// TIA Portal project "UploadAG314C_tia" (V15)

(* hardware
DEVICE "SIMATIC 300(1)"  S7-300 station
   slot 0: "Rack 0"  Rail  6ES7 390-1***0-0AA0
   slot 2: "CPU 314C-2 DP"  CPU 314C-2 DP  6ES7 314-6CG03-0AB0  V2.6
      slot 0: "MPI interface_1"  X1
      slot 1: "DP interface_1"  X2
      slot 2: "DI 24/DO 16_1"  DI24/DO16
      slot 3: "AI 5/AO 2_1"  AI5/AO2
      slot 4: "Count_1"  Counter
      slot 5: "Positioning_1"  Positioning
DEVICE "Test_Pump"  TP1200 Comfort
   slot 0: "Test_Pump"  TP1200 Comfort  6AV2 124-0MC01-0AX0  14.0.1.0
   slot 1: "HMI_RT_2"  TP1200 Comfort  6AV2 124-0MC01-0AX0  14.0.1.0
   slot 5: "Test_Pump._CP_1"  PROFINET Interface  14.0.1.0
      slot 1: "PROFINET Interface_1"  PROFINET Interface
         slot 1: "Port_1"  Port
         slot 2: "Port_2"  Port
   slot 7: "Test_Pump.I/DP_CP_1"  MPI/DP Interface  14.0.1.0
*)

// ===== PLC "CPU 314C-2 DP"  CPU 314C-2 DP =====
// protected blocks, not shown: "CONT_C_LF"

VAR_GLOBAL   // PLC tag table "Default tag table"
   "Tag_5" AT %M40.0 : Bool;
   "Tag_6" AT %M30.0 : Bool;
   "Tag_7" AT %M30.3 : Bool;
   "Tag_8" AT %M30.6 : Bool;
   "Tag_9" AT %M30.4 : Bool;
   "Tag_10" AT %M30.7 : Bool;
   "Tag_11" AT %M33.3 : Bool;
   "Tag_12" AT %M33.6 : Bool;
   "Tag_13" AT %M33.4 : Bool;
   "Tag_14" AT %M33.7 : Bool;
   "Tag_15" AT %I126.0 : Bool;
   "Tag_16" AT %M70.1 : Bool;
   "Tag_17" AT %I126.1 : Bool;
   "Tag_18" AT %M70.0 : Bool;
   "Tag_19" AT %I126.2 : Bool;
   "Tag_20" AT %I126.3 : Bool;
   "Tag_21" AT %I126.5 : Bool;
   "Tag_22" AT %I126.6 : Bool;
   "Tag_23" AT %Q124.1 : Bool;
   "Tag_24" AT %Q124.0 : Bool;
   "Tag_25" AT %M30.1 : Bool;
   "Tag_26" AT %M31.0 : Bool;
   "Tag_27" AT %T40 : Timer;
   "Tag_28" AT %Q124.2 : Bool;
   "Tag_29" AT %MD210 : DWord;
   "Tag_30" AT %MW212 : Word;
   "samplingTimer_1" AT %T190 : Timer;
   "samplingTimer_2" AT %T191 : Timer;
   "Tag_31" AT %M0.0 : Bool;
   "Tag_32" AT %T192 : Timer;
   "Speed" AT %MW4 : Int;
END_VAR

VAR_GLOBAL   // PLC tag table "STEP7 classic symbols"
   "Tag_1" AT %AW752 : Word;
   "Tag_2" AT %EW752 : Int;
   "Tag_3" AT %EW760 : Word;
   "Tag_4" AT %MD20 : DInt;
END_VAR

DATA_BLOCK "DB3"   // DB3
{ S7_Optimized_Access := 'FALSE' }
VERSION : 0.1
   VAR
      STAT0 : Word := WORD#16#0001;
      STAT1 : Word;
      STAT2 : Word := WORD#16#0009;
      STAT3 : Word := WORD#16#0003;
      STAT4 : Word := WORD#16#0027;
      STAT5 : Word := WORD#16#1456;
      STAT6 : Word;
      STAT7 : Word;
      STAT8 : Word;
      STAT9 : Word;
      STAT10 : Word;
      STAT11 : Word;
      STAT12 : Word;
      STAT13 : Word;
      STAT14 : Word;
      STAT15 : Word;
      STAT16 : Word;
      STAT17 : Word;
      STAT18 : Word;
      STAT19 : Word;
      STAT20 : Word;
   END_VAR
BEGIN
END_DATA_BLOCK

DATA_BLOCK "DB5"   // DB5
{ S7_Optimized_Access := 'FALSE' }
VERSION : 0.1
   VAR
      STAT0 : Word;
      STAT1 : Word := WORD#16#0400;
      STAT2 : Word;
      STAT3 : Word := WORD#16#0001;
      STAT4 : Word := WORD#16#0001;
      STAT5 : Word := WORD#16#0020;
      STAT6 : Word;
      STAT7 : Word;
      STAT8 : Word;
      STAT9 : Word;
      STAT10 : Word;
      STAT11 : Word;
      STAT12 : Word;
      STAT13 : Word;
      STAT14 : Word;
      STAT15 : Word;
      STAT16 : Word;
      STAT17 : Word;
      STAT18 : Word;
      STAT19 : Word;
      STAT20 : Word;
   END_VAR
BEGIN
END_DATA_BLOCK

DATA_BLOCK "DB12"   // DB12
{ S7_Optimized_Access := 'FALSE' }
VERSION : 0.1
   VAR
      STAT0 : Int;
      STAT1 : Int;
      STAT2 : Int := 250;
      STAT3 : Int := 336;
      STAT4 : DInt;
      STAT5 : DInt;
      STAT6 : DInt;
      STAT7 : DInt;
      STAT8 : DInt;
      STAT9 : DInt;
      STAT10 : DInt;
   END_VAR
BEGIN
END_DATA_BLOCK

DATA_BLOCK "DB13"   // DB13
{ S7_Optimized_Access := 'FALSE' }
VERSION : 0.1
   VAR
      STAT0 : Real;
      STAT1 : Real;
      STAT2 : Real;
      STAT3 : Real;
      STAT4 : Real;
      STAT5 : Real;
      STAT6 : Real;
      STAT7 : Real;
   END_VAR
BEGIN
END_DATA_BLOCK

DATA_BLOCK "DB14"   // DB14
{ S7_Optimized_Access := 'FALSE' }
VERSION : 0.1
   VAR
      STAT0 : Int;
      STAT1 : Int;
      STAT2 : DInt;
      STAT3 : DInt;
      STAT4 : DInt;
      STAT5 : Int;
      STAT6 : Int;
      STAT7 : Int := 410;
      STAT8 : Int;
      STAT9 : DInt;
      STAT10 : DInt;
      STAT11 : DInt;
      STAT12 : Int := 6800;
      STAT13 : Int;
      STAT14 : DInt;
      STAT15 : DInt;
      STAT16 : DInt;
      STAT17 : DInt;
      STAT18 : Real;
      STAT19 : Real;
      STAT20 : DInt;
      STAT21 : DInt := DINT#98300;
      STAT22 : Real;
      STAT23 : Real;
      STAT24 : Real;
   END_VAR
BEGIN
END_DATA_BLOCK

DATA_BLOCK "DB16"   // DB16
{ S7_Optimized_Access := 'FALSE' }
VERSION : 0.1
   VAR
      STAT0 : Int;
      STAT1 : String[10];
      STAT2 : DInt;
      STAT3 : DInt;
      STAT4 : DInt;
      STAT5 : DInt := DINT#750;
      STAT6 : DInt;
      STAT7 : DInt;
      STAT8 : DInt;
      STAT9 : DInt;
      STAT10 : DInt;
      STAT11 : DInt;
      STAT12 : DInt;
      STAT13 : Int;
      STAT14 : Int := 1;
      STAT15 : String[10];
      STAT16 : DInt;
      STAT17 : DInt;
      STAT18 : DInt;
      STAT19 : DInt;
      STAT20 : DInt;
      STAT21 : DInt;
      STAT22 : DInt;
      STAT23 : DInt;
      STAT24 : DInt;
      STAT25 : DInt;
      STAT26 : DInt;
      STAT27 : Int;
      STAT28 : Int := 2;
      STAT29 : String[10];
      STAT30 : DInt;
      STAT31 : DInt;
      STAT32 : DInt;
      STAT33 : DInt;
      STAT34 : DInt;
      STAT35 : DInt;
      STAT36 : DInt;
      STAT37 : DInt;
      STAT38 : DInt;
      STAT39 : DInt;
      STAT40 : DInt;
      STAT41 : Int;
      STAT42 : Int := 3;
      STAT43 : String[10];
      STAT44 : DInt;
      STAT45 : DInt;
      STAT46 : DInt;
      STAT47 : DInt;
      STAT48 : DInt;
      STAT49 : DInt;
      STAT50 : DInt;
      STAT51 : DInt;
      STAT52 : DInt;
      STAT53 : DInt;
      STAT54 : DInt;
      STAT55 : Int;
      STAT56 : Int := 4;
      STAT57 : String[10];
      STAT58 : DInt;
      STAT59 : DInt;
      STAT60 : DInt;
      STAT61 : DInt;
      STAT62 : DInt;
      STAT63 : DInt;
      STAT64 : DInt;
      STAT65 : DInt;
      STAT66 : DInt;
      STAT67 : DInt;
      STAT68 : DInt;
      STAT69 : Int;
      STAT70 : Int := 5;
      STAT71 : String[10];
      STAT72 : DInt;
      STAT73 : DInt;
      STAT74 : DInt;
      STAT75 : DInt;
      STAT76 : DInt;
      STAT77 : DInt;
      STAT78 : DInt;
      STAT79 : DInt;
      STAT80 : DInt;
      STAT81 : DInt;
      STAT82 : DInt;
      STAT83 : Int;
      STAT84 : Int := 6;
      STAT85 : String[10];
      STAT86 : DInt;
      STAT87 : DInt;
      STAT88 : DInt;
      STAT89 : DInt;
      STAT90 : DInt;
      STAT91 : DInt;
      STAT92 : DInt;
      STAT93 : DInt;
      STAT94 : DInt;
      STAT95 : DInt;
      STAT96 : DInt;
      STAT97 : Int;
      STAT98 : Int := 7;
      STAT99 : String[10];
      STAT100 : DInt;
      STAT101 : DInt;
      STAT102 : DInt;
      STAT103 : DInt;
      STAT104 : DInt;
      STAT105 : DInt;
      STAT106 : DInt;
      STAT107 : DInt;
      STAT108 : DInt;
      STAT109 : DInt;
      STAT110 : DInt;
      STAT111 : Int;
      STAT112 : Int := 8;
      STAT113 : String[10];
      STAT114 : DInt;
      STAT115 : DInt;
      STAT116 : DInt;
      STAT117 : DInt;
      STAT118 : DInt;
      STAT119 : DInt;
      STAT120 : DInt;
      STAT121 : DInt;
      STAT122 : DInt;
      STAT123 : DInt;
      STAT124 : DInt;
      STAT125 : Int;
      STAT126 : Int := 9;
      STAT127 : String[10];
      STAT128 : DInt;
      STAT129 : DInt;
      STAT130 : DInt;
      STAT131 : DInt;
      STAT132 : DInt;
      STAT133 : DInt;
      STAT134 : DInt;
      STAT135 : DInt;
      STAT136 : DInt;
      STAT137 : DInt;
      STAT138 : DInt;
      STAT139 : Int;
      STAT140 : Int := 10;
      STAT141 : String[10];
      STAT142 : DInt;
      STAT143 : DInt;
      STAT144 : DInt;
      STAT145 : DInt;
      STAT146 : DInt;
      STAT147 : DInt;
      STAT148 : DInt;
      STAT149 : DInt;
      STAT150 : DInt;
      STAT151 : DInt;
      STAT152 : DInt;
      STAT153 : Int;
      STAT154 : Int := 11;
      STAT155 : String[10];
      STAT156 : DInt;
      STAT157 : DInt;
      STAT158 : DInt;
      STAT159 : DInt;
      STAT160 : DInt;
      STAT161 : DInt;
      STAT162 : DInt;
      STAT163 : DInt;
      STAT164 : DInt;
      STAT165 : DInt;
      STAT166 : DInt;
      STAT167 : Int;
      STAT168 : Int := 12;
      STAT169 : String[10];
      STAT170 : DInt;
      STAT171 : DInt;
      STAT172 : DInt;
      STAT173 : DInt;
      STAT174 : DInt;
      STAT175 : DInt;
      STAT176 : DInt;
      STAT177 : DInt;
      STAT178 : DInt;
      STAT179 : DInt;
      STAT180 : DInt;
      STAT181 : Int;
      STAT182 : Int := 13;
      STAT183 : String[10];
      STAT184 : DInt;
      STAT185 : DInt;
      STAT186 : DInt;
      STAT187 : DInt;
      STAT188 : DInt;
      STAT189 : DInt;
      STAT190 : DInt;
      STAT191 : DInt;
      STAT192 : DInt;
      STAT193 : DInt;
      STAT194 : DInt;
      STAT195 : Int;
      STAT196 : Int := 14;
      STAT197 : String[10];
      STAT198 : DInt;
      STAT199 : DInt;
      STAT200 : DInt;
      STAT201 : DInt;
      STAT202 : DInt;
      STAT203 : DInt;
      STAT204 : DInt;
      STAT205 : DInt;
      STAT206 : DInt;
      STAT207 : DInt;
      STAT208 : DInt;
      STAT209 : Int;
      STAT210 : Int := 15;
      STAT211 : String[10];
      STAT212 : DInt;
      STAT213 : DInt;
      STAT214 : DInt;
      STAT215 : DInt;
      STAT216 : DInt;
      STAT217 : DInt;
      STAT218 : DInt;
      STAT219 : DInt;
      STAT220 : DInt;
      STAT221 : DInt;
      STAT222 : DInt;
      STAT223 : Int;
      STAT224 : Int := 16;
      STAT225 : String[10];
      STAT226 : DInt;
      STAT227 : DInt;
      STAT228 : DInt;
      STAT229 : DInt;
      STAT230 : DInt;
      STAT231 : DInt;
      STAT232 : DInt;
      STAT233 : DInt;
      STAT234 : DInt;
      STAT235 : DInt;
      STAT236 : DInt;
      STAT237 : Int;
      STAT238 : Int := 17;
      STAT239 : String[10];
      STAT240 : DInt;
      STAT241 : DInt;
      STAT242 : DInt;
      STAT243 : DInt;
      STAT244 : DInt;
      STAT245 : DInt;
      STAT246 : DInt;
      STAT247 : DInt;
      STAT248 : DInt;
      STAT249 : DInt;
      STAT250 : DInt;
      STAT251 : Int;
      STAT252 : Int := 18;
      STAT253 : String[10];
      STAT254 : DInt;
      STAT255 : DInt;
      STAT256 : DInt;
      STAT257 : DInt;
      STAT258 : DInt;
      STAT259 : DInt;
      STAT260 : DInt;
      STAT261 : DInt;
      STAT262 : DInt;
      STAT263 : DInt;
      STAT264 : DInt;
      STAT265 : Int;
      STAT266 : Int := 19;
      STAT267 : String[10];
      STAT268 : DInt;
      STAT269 : DInt;
      STAT270 : DInt;
      STAT271 : DInt;
      STAT272 : DInt;
      STAT273 : DInt;
      STAT274 : DInt;
      STAT275 : DInt;
      STAT276 : DInt;
      STAT277 : DInt;
      STAT278 : DInt;
      STAT279 : Int;
      STAT280 : Int := 20;
      STAT281 : String[10];
      STAT282 : DInt;
      STAT283 : DInt;
      STAT284 : DInt;
      STAT285 : DInt;
      STAT286 : DInt;
      STAT287 : DInt;
      STAT288 : DInt;
      STAT289 : DInt;
      STAT290 : DInt;
      STAT291 : DInt;
      STAT292 : DInt;
      STAT293 : Int;
      STAT294 : Int := 21;
      STAT295 : String[10];
      STAT296 : DInt;
      STAT297 : DInt;
      STAT298 : DInt;
      STAT299 : DInt;
      STAT300 : DInt;
      STAT301 : DInt;
      STAT302 : DInt;
      STAT303 : DInt;
      STAT304 : DInt;
      STAT305 : DInt;
      STAT306 : DInt;
      STAT307 : Int;
      STAT308 : Int := 22;
      STAT309 : String[10];
      STAT310 : DInt;
      STAT311 : DInt;
      STAT312 : DInt;
      STAT313 : DInt;
      STAT314 : DInt;
      STAT315 : DInt;
      STAT316 : DInt;
      STAT317 : DInt;
      STAT318 : DInt;
      STAT319 : DInt;
      STAT320 : DInt;
      STAT321 : Int;
      STAT322 : Int := 23;
      STAT323 : String[10];
      STAT324 : DInt;
      STAT325 : DInt;
      STAT326 : DInt;
      STAT327 : DInt;
      STAT328 : DInt;
      STAT329 : DInt;
      STAT330 : DInt;
      STAT331 : DInt;
      STAT332 : DInt;
      STAT333 : DInt;
      STAT334 : DInt;
      STAT335 : Int;
      STAT336 : Int := 24;
      STAT337 : String[10];
      STAT338 : DInt;
      STAT339 : DInt;
      STAT340 : DInt;
      STAT341 : DInt;
      STAT342 : DInt;
      STAT343 : DInt;
      STAT344 : DInt;
      STAT345 : DInt;
      STAT346 : DInt;
      STAT347 : DInt;
      STAT348 : DInt;
      STAT349 : Int;
      STAT350 : Int := 25;
      STAT351 : String[10];
      STAT352 : DInt;
      STAT353 : DInt;
      STAT354 : DInt;
      STAT355 : DInt;
      STAT356 : DInt;
      STAT357 : DInt;
      STAT358 : DInt;
      STAT359 : DInt;
      STAT360 : DInt;
      STAT361 : DInt;
      STAT362 : DInt;
      STAT363 : Int;
      STAT364 : Int := 26;
      STAT365 : String[10];
      STAT366 : DInt;
      STAT367 : DInt;
      STAT368 : DInt;
      STAT369 : DInt;
      STAT370 : DInt;
      STAT371 : DInt;
      STAT372 : DInt;
      STAT373 : DInt;
      STAT374 : DInt;
      STAT375 : DInt;
      STAT376 : DInt;
      STAT377 : Int;
      STAT378 : Int := 27;
      STAT379 : String[10];
      STAT380 : DInt;
      STAT381 : DInt;
      STAT382 : DInt;
      STAT383 : DInt;
      STAT384 : DInt;
      STAT385 : DInt;
      STAT386 : DInt;
      STAT387 : DInt;
      STAT388 : DInt;
      STAT389 : DInt;
      STAT390 : DInt;
      STAT391 : Int;
      STAT392 : Int := 28;
      STAT393 : String[10];
      STAT394 : DInt;
      STAT395 : DInt;
      STAT396 : DInt;
      STAT397 : DInt;
      STAT398 : DInt;
      STAT399 : DInt;
      STAT400 : DInt;
      STAT401 : DInt;
      STAT402 : DInt;
      STAT403 : DInt;
      STAT404 : DInt;
      STAT405 : Int;
      STAT406 : Int := 29;
      STAT407 : String[10];
      STAT408 : DInt;
      STAT409 : DInt;
      STAT410 : DInt;
      STAT411 : DInt;
      STAT412 : DInt;
      STAT413 : DInt;
      STAT414 : DInt;
      STAT415 : DInt;
      STAT416 : DInt;
      STAT417 : DInt;
      STAT418 : DInt;
      STAT419 : Int;
      STAT420 : Int := 30;
      STAT421 : String[10];
      STAT422 : DInt;
      STAT423 : DInt;
      STAT424 : DInt;
      STAT425 : DInt;
      STAT426 : DInt;
      STAT427 : DInt;
      STAT428 : DInt;
      STAT429 : DInt;
      STAT430 : DInt;
      STAT431 : DInt;
      STAT432 : DInt;
      STAT433 : Int;
      STAT434 : Int := 31;
      STAT435 : String[10];
      STAT436 : DInt;
      STAT437 : DInt;
      STAT438 : DInt;
      STAT439 : DInt;
      STAT440 : DInt;
      STAT441 : DInt;
      STAT442 : DInt;
      STAT443 : DInt;
      STAT444 : DInt;
      STAT445 : DInt;
      STAT446 : DInt;
      STAT447 : Int;
      STAT448 : Int := 32;
      STAT449 : String[10];
      STAT450 : DInt;
      STAT451 : DInt;
      STAT452 : DInt;
      STAT453 : DInt;
      STAT454 : DInt;
      STAT455 : DInt;
      STAT456 : DInt;
      STAT457 : DInt;
      STAT458 : DInt;
      STAT459 : DInt;
      STAT460 : DInt;
      STAT461 : Int;
      STAT462 : Int := 33;
      STAT463 : String[10];
      STAT464 : DInt;
      STAT465 : DInt;
      STAT466 : DInt;
      STAT467 : DInt;
      STAT468 : DInt;
      STAT469 : DInt;
      STAT470 : DInt;
      STAT471 : DInt;
      STAT472 : DInt;
      STAT473 : DInt;
      STAT474 : DInt;
      STAT475 : Int;
      STAT476 : Int := 34;
      STAT477 : String[10];
      STAT478 : DInt;
      STAT479 : DInt;
      STAT480 : DInt;
      STAT481 : DInt;
      STAT482 : DInt;
      STAT483 : DInt;
      STAT484 : DInt;
      STAT485 : DInt;
      STAT486 : DInt;
      STAT487 : DInt;
      STAT488 : DInt;
      STAT489 : Int;
      STAT490 : Int := 35;
      STAT491 : String[10];
      STAT492 : DInt;
      STAT493 : DInt;
      STAT494 : DInt;
      STAT495 : DInt;
      STAT496 : DInt;
      STAT497 : DInt;
      STAT498 : DInt;
      STAT499 : DInt;
      STAT500 : DInt;
      STAT501 : DInt;
      STAT502 : DInt;
      STAT503 : Int;
      STAT504 : Int := 36;
      STAT505 : String[10];
      STAT506 : DInt;
      STAT507 : DInt;
      STAT508 : DInt;
      STAT509 : DInt;
      STAT510 : DInt;
      STAT511 : DInt;
      STAT512 : DInt;
      STAT513 : DInt;
      STAT514 : DInt;
      STAT515 : DInt;
      STAT516 : DInt;
      STAT517 : Int;
      STAT518 : Int := 37;
      STAT519 : String[10];
      STAT520 : DInt;
      STAT521 : DInt;
      STAT522 : DInt;
      STAT523 : DInt;
      STAT524 : DInt;
      STAT525 : DInt;
      STAT526 : DInt;
      STAT527 : DInt;
      STAT528 : DInt;
      STAT529 : DInt;
      STAT530 : DInt;
      STAT531 : Int;
      STAT532 : Int := 38;
      STAT533 : String[10];
      STAT534 : DInt;
      STAT535 : DInt;
      STAT536 : DInt;
      STAT537 : DInt;
      STAT538 : DInt;
      STAT539 : DInt;
      STAT540 : DInt;
      STAT541 : DInt;
      STAT542 : DInt;
      STAT543 : DInt;
      STAT544 : DInt;
      STAT545 : Int;
      STAT546 : Int := 39;
      STAT547 : String[10];
      STAT548 : DInt;
      STAT549 : DInt;
      STAT550 : DInt;
      STAT551 : DInt;
      STAT552 : DInt;
      STAT553 : DInt;
      STAT554 : DInt;
      STAT555 : DInt;
      STAT556 : DInt;
      STAT557 : DInt;
      STAT558 : DInt;
      STAT559 : Int;
      STAT560 : Int := 40;
      STAT561 : String[10];
      STAT562 : DInt;
      STAT563 : DInt;
      STAT564 : DInt;
      STAT565 : DInt;
      STAT566 : DInt;
      STAT567 : DInt;
      STAT568 : DInt;
      STAT569 : DInt;
      STAT570 : DInt;
      STAT571 : DInt;
      STAT572 : DInt;
      STAT573 : Int;
      STAT574 : Int := 41;
      STAT575 : String[10];
      STAT576 : DInt;
      STAT577 : DInt;
      STAT578 : DInt;
      STAT579 : DInt;
      STAT580 : DInt;
      STAT581 : DInt;
      STAT582 : DInt;
      STAT583 : DInt;
      STAT584 : DInt;
      STAT585 : DInt;
      STAT586 : DInt;
      STAT587 : Int;
      STAT588 : Int := 42;
      STAT589 : String[10];
      STAT590 : DInt;
      STAT591 : DInt;
      STAT592 : DInt;
      STAT593 : DInt;
      STAT594 : DInt;
      STAT595 : DInt;
      STAT596 : DInt;
      STAT597 : DInt;
      STAT598 : DInt;
      STAT599 : DInt;
      STAT600 : DInt;
      STAT601 : Int;
      STAT602 : Int := 43;
      STAT603 : String[10];
      STAT604 : DInt;
      STAT605 : DInt;
      STAT606 : DInt;
      STAT607 : DInt;
      STAT608 : DInt;
      STAT609 : DInt;
      STAT610 : DInt;
      STAT611 : DInt;
      STAT612 : DInt;
      STAT613 : DInt;
      STAT614 : DInt;
      STAT615 : Int;
      STAT616 : Int := 44;
      STAT617 : String[10];
      STAT618 : DInt;
      STAT619 : DInt;
      STAT620 : DInt;
      STAT621 : DInt;
      STAT622 : DInt;
      STAT623 : DInt;
      STAT624 : DInt;
      STAT625 : DInt;
      STAT626 : DInt;
      STAT627 : DInt;
      STAT628 : DInt;
      STAT629 : Int;
      STAT630 : Int := 45;
      STAT631 : String[10];
      STAT632 : DInt;
      STAT633 : DInt;
      STAT634 : DInt;
      STAT635 : DInt;
      STAT636 : DInt;
      STAT637 : DInt;
      STAT638 : DInt;
      STAT639 : DInt;
      STAT640 : DInt;
      STAT641 : DInt;
      STAT642 : DInt;
      STAT643 : Int;
      STAT644 : Int := 46;
      STAT645 : String[10];
      STAT646 : DInt;
      STAT647 : DInt;
      STAT648 : DInt;
      STAT649 : DInt;
      STAT650 : DInt;
      STAT651 : DInt;
      STAT652 : DInt;
      STAT653 : DInt;
      STAT654 : DInt;
      STAT655 : DInt;
      STAT656 : DInt;
      STAT657 : Int;
      STAT658 : Int := 47;
      STAT659 : String[10];
      STAT660 : DInt;
      STAT661 : DInt;
      STAT662 : DInt;
      STAT663 : DInt;
      STAT664 : DInt;
      STAT665 : DInt;
      STAT666 : DInt;
      STAT667 : DInt;
      STAT668 : DInt;
      STAT669 : DInt;
      STAT670 : DInt;
      STAT671 : Int;
      STAT672 : Int := 48;
      STAT673 : String[10];
      STAT674 : DInt;
      STAT675 : DInt;
      STAT676 : DInt;
      STAT677 : DInt;
      STAT678 : DInt;
      STAT679 : DInt;
      STAT680 : DInt;
      STAT681 : DInt;
      STAT682 : DInt;
      STAT683 : DInt;
      STAT684 : DInt;
      STAT685 : Int;
      STAT686 : Int := 49;
      STAT687 : String[10];
      STAT688 : DInt;
      STAT689 : DInt;
      STAT690 : DInt;
      STAT691 : DInt;
      STAT692 : DInt;
      STAT693 : DInt;
      STAT694 : DInt;
      STAT695 : DInt;
      STAT696 : DInt;
      STAT697 : DInt;
      STAT698 : DInt;
      STAT699 : Int;
      STAT700 : Int := 50;
      STAT701 : String[10];
      STAT702 : DInt;
      STAT703 : DInt;
      STAT704 : DInt;
      STAT705 : DInt;
      STAT706 : DInt;
      STAT707 : DInt;
      STAT708 : DInt;
      STAT709 : DInt;
      STAT710 : DInt;
      STAT711 : DInt;
      STAT712 : DInt;
      STAT713 : Int;
      STAT714 : Int := 51;
      STAT715 : String[10];
      STAT716 : DInt;
      STAT717 : DInt;
      STAT718 : DInt;
      STAT719 : DInt;
      STAT720 : DInt;
      STAT721 : DInt;
      STAT722 : DInt;
      STAT723 : DInt;
      STAT724 : DInt;
      STAT725 : DInt;
      STAT726 : DInt;
      STAT727 : Int;
      STAT728 : Int := 52;
      STAT729 : String[10];
      STAT730 : DInt;
      STAT731 : DInt;
      STAT732 : DInt;
      STAT733 : DInt;
      STAT734 : DInt;
      STAT735 : DInt;
      STAT736 : DInt;
      STAT737 : DInt;
      STAT738 : DInt;
      STAT739 : DInt;
      STAT740 : DInt;
      STAT741 : Int;
      STAT742 : Int := 53;
      STAT743 : String[10];
      STAT744 : DInt;
      STAT745 : DInt;
      STAT746 : DInt;
      STAT747 : DInt;
      STAT748 : DInt;
      STAT749 : DInt;
      STAT750 : DInt;
      STAT751 : DInt;
      STAT752 : DInt;
      STAT753 : DInt;
      STAT754 : DInt;
      STAT755 : Int;
      STAT756 : Int := 54;
      STAT757 : String[10];
      STAT758 : DInt;
      STAT759 : DInt;
      STAT760 : DInt;
      STAT761 : DInt;
      STAT762 : DInt;
      STAT763 : DInt;
      STAT764 : DInt;
      STAT765 : DInt;
      STAT766 : DInt;
      STAT767 : DInt;
      STAT768 : DInt;
      STAT769 : Int;
      STAT770 : Int := 55;
      STAT771 : String[10];
      STAT772 : DInt;
      STAT773 : DInt;
      STAT774 : DInt;
      STAT775 : DInt;
      STAT776 : DInt;
      STAT777 : DInt;
      STAT778 : DInt;
      STAT779 : DInt;
      STAT780 : DInt;
      STAT781 : DInt;
      STAT782 : DInt;
      STAT783 : Int;
      STAT784 : Int := 56;
      STAT785 : String[10];
      STAT786 : DInt;
      STAT787 : DInt;
      STAT788 : DInt;
      STAT789 : DInt;
      STAT790 : DInt;
      STAT791 : DInt;
      STAT792 : DInt;
      STAT793 : DInt;
      STAT794 : DInt;
      STAT795 : DInt;
      STAT796 : DInt;
      STAT797 : Int;
      STAT798 : Int := 57;
      STAT799 : String[10];
      STAT800 : DInt;
      STAT801 : DInt;
      STAT802 : DInt;
      STAT803 : DInt;
      STAT804 : DInt;
      STAT805 : DInt;
      STAT806 : DInt;
      STAT807 : DInt;
      STAT808 : DInt;
      STAT809 : DInt;
      STAT810 : DInt;
      STAT811 : Int;
      STAT812 : Int := 58;
      STAT813 : String[10];
      STAT814 : DInt;
      STAT815 : DInt;
      STAT816 : DInt;
      STAT817 : DInt;
      STAT818 : DInt;
      STAT819 : DInt;
      STAT820 : DInt;
      STAT821 : DInt;
      STAT822 : DInt;
      STAT823 : DInt;
      STAT824 : DInt;
      STAT825 : Int;
      STAT826 : Int := 59;
      STAT827 : String[10];
      STAT828 : DInt;
      STAT829 : DInt;
      STAT830 : DInt;
      STAT831 : DInt;
      STAT832 : DInt;
      STAT833 : DInt;
      STAT834 : DInt;
      STAT835 : DInt;
      STAT836 : DInt;
      STAT837 : DInt;
      STAT838 : DInt;
      STAT839 : Int;
      STAT840 : Int := 60;
      STAT841 : String[10];
      STAT842 : DInt;
      STAT843 : DInt;
      STAT844 : DInt;
      STAT845 : DInt;
      STAT846 : DInt;
      STAT847 : DInt;
      STAT848 : DInt;
      STAT849 : DInt;
      STAT850 : DInt;
      STAT851 : DInt;
      STAT852 : DInt;
      STAT853 : Int;
      STAT854 : Int := 61;
      STAT855 : String[10];
      STAT856 : DInt;
      STAT857 : DInt;
      STAT858 : DInt;
      STAT859 : DInt;
      STAT860 : DInt;
      STAT861 : DInt;
      STAT862 : DInt;
      STAT863 : DInt;
      STAT864 : DInt;
      STAT865 : DInt;
      STAT866 : DInt;
      STAT867 : Int;
      STAT868 : Int := 62;
      STAT869 : String[10];
      STAT870 : DInt;
      STAT871 : DInt;
      STAT872 : DInt;
      STAT873 : DInt;
      STAT874 : DInt;
      STAT875 : DInt;
      STAT876 : DInt;
      STAT877 : DInt;
      STAT878 : DInt;
      STAT879 : DInt;
      STAT880 : DInt;
      STAT881 : Int;
      STAT882 : Int := 63;
      STAT883 : String[10];
      STAT884 : DInt;
      STAT885 : DInt;
      STAT886 : DInt;
      STAT887 : DInt;
      STAT888 : DInt;
      STAT889 : DInt;
      STAT890 : DInt;
      STAT891 : DInt;
      STAT892 : DInt;
      STAT893 : DInt;
      STAT894 : DInt;
      STAT895 : Int;
      STAT896 : Int := 64;
      STAT897 : String[10];
      STAT898 : DInt;
      STAT899 : DInt;
      STAT900 : DInt;
      STAT901 : DInt;
      STAT902 : DInt;
      STAT903 : DInt;
      STAT904 : DInt;
      STAT905 : DInt;
      STAT906 : DInt;
      STAT907 : DInt;
      STAT908 : DInt;
      STAT909 : Int;
      STAT910 : Int := 65;
      STAT911 : String[10];
      STAT912 : DInt;
      STAT913 : DInt;
      STAT914 : DInt;
      STAT915 : DInt;
      STAT916 : DInt;
      STAT917 : DInt;
      STAT918 : DInt;
      STAT919 : DInt;
      STAT920 : DInt;
      STAT921 : DInt;
      STAT922 : DInt;
      STAT923 : Int;
      STAT924 : Int := 66;
      STAT925 : String[10];
      STAT926 : DInt;
      STAT927 : DInt;
      STAT928 : DInt;
      STAT929 : DInt;
      STAT930 : DInt;
      STAT931 : DInt;
      STAT932 : DInt;
      STAT933 : DInt;
      STAT934 : DInt;
      STAT935 : DInt;
      STAT936 : DInt;
      STAT937 : Int;
      STAT938 : Int := 67;
      STAT939 : String[10];
      STAT940 : DInt;
      STAT941 : DInt;
      STAT942 : DInt;
      STAT943 : DInt;
      STAT944 : DInt;
      STAT945 : DInt;
      STAT946 : DInt;
      STAT947 : DInt;
      STAT948 : DInt;
      STAT949 : DInt;
      STAT950 : DInt;
      STAT951 : Int;
      STAT952 : Int := 68;
      STAT953 : String[10];
      STAT954 : DInt;
      STAT955 : DInt;
      STAT956 : DInt;
      STAT957 : DInt;
      STAT958 : DInt;
      STAT959 : DInt;
      STAT960 : DInt;
      STAT961 : DInt;
      STAT962 : DInt;
      STAT963 : DInt;
      STAT964 : DInt;
      STAT965 : Int;
      STAT966 : Int := 69;
      STAT967 : String[10];
      STAT968 : DInt;
      STAT969 : DInt;
      STAT970 : DInt;
      STAT971 : DInt;
      STAT972 : DInt;
      STAT973 : DInt;
      STAT974 : DInt;
      STAT975 : DInt;
      STAT976 : DInt;
      STAT977 : DInt;
      STAT978 : DInt;
      STAT979 : Int;
      STAT980 : Int := 70;
      STAT981 : String[10];
      STAT982 : DInt;
      STAT983 : DInt;
      STAT984 : DInt;
      STAT985 : DInt;
      STAT986 : DInt;
      STAT987 : DInt;
      STAT988 : DInt;
      STAT989 : DInt;
      STAT990 : DInt;
      STAT991 : DInt;
      STAT992 : DInt;
      STAT993 : Int;
      STAT994 : Int := 71;
      STAT995 : String[10];
      STAT996 : DInt;
      STAT997 : DInt;
      STAT998 : DInt;
      STAT999 : DInt;
      STAT1000 : DInt;
      STAT1001 : DInt;
      STAT1002 : DInt;
      STAT1003 : DInt;
      STAT1004 : DInt;
      STAT1005 : DInt;
      STAT1006 : DInt;
      STAT1007 : Int;
      STAT1008 : Int := 72;
      STAT1009 : String[10];
      STAT1010 : DInt;
      STAT1011 : DInt;
      STAT1012 : DInt;
      STAT1013 : DInt;
      STAT1014 : DInt;
      STAT1015 : DInt;
      STAT1016 : DInt;
      STAT1017 : DInt;
      STAT1018 : DInt;
      STAT1019 : DInt;
      STAT1020 : DInt;
      STAT1021 : Int;
      STAT1022 : Int := 73;
      STAT1023 : String[10];
      STAT1024 : DInt;
      STAT1025 : DInt;
      STAT1026 : DInt;
      STAT1027 : DInt;
      STAT1028 : DInt;
      STAT1029 : DInt;
      STAT1030 : DInt;
      STAT1031 : DInt;
      STAT1032 : DInt;
      STAT1033 : DInt;
      STAT1034 : DInt;
      STAT1035 : Int;
      STAT1036 : Int := 74;
      STAT1037 : String[10];
      STAT1038 : DInt;
      STAT1039 : DInt;
      STAT1040 : DInt;
      STAT1041 : DInt;
      STAT1042 : DInt;
      STAT1043 : DInt;
      STAT1044 : DInt;
      STAT1045 : DInt;
      STAT1046 : DInt;
      STAT1047 : DInt;
      STAT1048 : DInt;
      STAT1049 : Int;
      STAT1050 : Int := 75;
      STAT1051 : String[10];
      STAT1052 : DInt;
      STAT1053 : DInt;
      STAT1054 : DInt;
      STAT1055 : DInt;
      STAT1056 : DInt;
      STAT1057 : DInt;
      STAT1058 : DInt;
      STAT1059 : DInt;
      STAT1060 : DInt;
      STAT1061 : DInt;
      STAT1062 : DInt;
      STAT1063 : Int;
      STAT1064 : Int := 76;
      STAT1065 : String[10];
      STAT1066 : DInt;
      STAT1067 : DInt;
      STAT1068 : DInt;
      STAT1069 : DInt;
      STAT1070 : DInt;
      STAT1071 : DInt;
      STAT1072 : DInt;
      STAT1073 : DInt;
      STAT1074 : DInt;
      STAT1075 : DInt;
      STAT1076 : DInt;
      STAT1077 : Int;
      STAT1078 : Int := 77;
      STAT1079 : String[10];
      STAT1080 : DInt;
      STAT1081 : DInt;
      STAT1082 : DInt;
      STAT1083 : DInt;
      STAT1084 : DInt;
      STAT1085 : DInt;
      STAT1086 : DInt;
      STAT1087 : DInt;
      STAT1088 : DInt;
      STAT1089 : DInt;
      STAT1090 : DInt;
      STAT1091 : Int;
      STAT1092 : Int := 78;
      STAT1093 : String[10];
      STAT1094 : DInt;
      STAT1095 : DInt;
      STAT1096 : DInt;
      STAT1097 : DInt;
      STAT1098 : DInt;
      STAT1099 : DInt;
      STAT1100 : DInt;
      STAT1101 : DInt;
      STAT1102 : DInt;
      STAT1103 : DInt;
      STAT1104 : DInt;
      STAT1105 : Int;
      STAT1106 : Int := 79;
      STAT1107 : String[10];
      STAT1108 : DInt;
      STAT1109 : DInt;
      STAT1110 : DInt;
      STAT1111 : DInt;
      STAT1112 : DInt;
      STAT1113 : DInt;
      STAT1114 : DInt;
      STAT1115 : DInt;
      STAT1116 : DInt;
      STAT1117 : DInt;
      STAT1118 : DInt;
      STAT1119 : Int;
      STAT1120 : Int := 80;
      STAT1121 : String[10];
      STAT1122 : DInt;
      STAT1123 : DInt;
      STAT1124 : DInt;
      STAT1125 : DInt;
      STAT1126 : DInt;
      STAT1127 : DInt;
      STAT1128 : DInt;
      STAT1129 : DInt;
      STAT1130 : DInt;
      STAT1131 : DInt;
      STAT1132 : DInt;
      STAT1133 : Int;
      STAT1134 : Int := 81;
      STAT1135 : String[10];
      STAT1136 : DInt;
      STAT1137 : DInt;
      STAT1138 : DInt;
      STAT1139 : DInt;
      STAT1140 : DInt;
      STAT1141 : DInt;
      STAT1142 : DInt;
      STAT1143 : DInt;
      STAT1144 : DInt;
      STAT1145 : DInt;
      STAT1146 : DInt;
      STAT1147 : Int;
      STAT1148 : Int := 82;
      STAT1149 : String[10];
      STAT1150 : DInt;
      STAT1151 : DInt;
      STAT1152 : DInt;
      STAT1153 : DInt;
      STAT1154 : DInt;
      STAT1155 : DInt;
      STAT1156 : DInt;
      STAT1157 : DInt;
      STAT1158 : DInt;
      STAT1159 : DInt;
      STAT1160 : DInt;
      STAT1161 : Int;
      STAT1162 : Int := 83;
      STAT1163 : String[10];
      STAT1164 : DInt;
      STAT1165 : DInt;
      STAT1166 : DInt;
      STAT1167 : DInt;
      STAT1168 : DInt;
      STAT1169 : DInt;
      STAT1170 : DInt;
      STAT1171 : DInt;
      STAT1172 : DInt;
      STAT1173 : DInt;
      STAT1174 : DInt;
      STAT1175 : Int;
      STAT1176 : Int := 84;
      STAT1177 : String[10];
      STAT1178 : DInt;
      STAT1179 : DInt;
      STAT1180 : DInt;
      STAT1181 : DInt;
      STAT1182 : DInt;
      STAT1183 : DInt;
      STAT1184 : DInt;
      STAT1185 : DInt;
      STAT1186 : DInt;
      STAT1187 : DInt;
      STAT1188 : DInt;
      STAT1189 : Int;
      STAT1190 : Int := 85;
      STAT1191 : String[10];
      STAT1192 : DInt;
      STAT1193 : DInt;
      STAT1194 : DInt;
      STAT1195 : DInt;
      STAT1196 : DInt;
      STAT1197 : DInt;
      STAT1198 : DInt;
      STAT1199 : DInt;
      STAT1200 : DInt;
      STAT1201 : DInt;
      STAT1202 : DInt;
      STAT1203 : Int;
      STAT1204 : Int := 86;
      STAT1205 : String[10];
      STAT1206 : DInt;
      STAT1207 : DInt;
      STAT1208 : DInt;
      STAT1209 : DInt;
      STAT1210 : DInt;
      STAT1211 : DInt;
      STAT1212 : DInt;
      STAT1213 : DInt;
      STAT1214 : DInt;
      STAT1215 : DInt;
      STAT1216 : DInt;
      STAT1217 : Int;
      STAT1218 : Int := 87;
      STAT1219 : String[10];
      STAT1220 : DInt;
      STAT1221 : DInt;
      STAT1222 : DInt;
      STAT1223 : DInt;
      STAT1224 : DInt;
      STAT1225 : DInt;
      STAT1226 : DInt;
      STAT1227 : DInt;
      STAT1228 : DInt;
      STAT1229 : DInt;
      STAT1230 : DInt;
      STAT1231 : Int;
      STAT1232 : Int := 88;
      STAT1233 : String[10];
      STAT1234 : DInt;
      STAT1235 : DInt;
      STAT1236 : DInt;
      STAT1237 : DInt;
      STAT1238 : DInt;
      STAT1239 : DInt;
      STAT1240 : DInt;
      STAT1241 : DInt;
      STAT1242 : DInt;
      STAT1243 : DInt;
      STAT1244 : DInt;
      STAT1245 : Int;
      STAT1246 : Int := 89;
      STAT1247 : String[10];
      STAT1248 : DInt;
      STAT1249 : DInt;
      STAT1250 : DInt;
      STAT1251 : DInt;
      STAT1252 : DInt;
      STAT1253 : DInt;
      STAT1254 : DInt;
      STAT1255 : DInt;
      STAT1256 : DInt;
      STAT1257 : DInt;
      STAT1258 : DInt;
      STAT1259 : Int;
      STAT1260 : Int := 90;
      STAT1261 : String[10];
      STAT1262 : DInt;
      STAT1263 : DInt;
      STAT1264 : DInt;
      STAT1265 : DInt;
      STAT1266 : DInt;
      STAT1267 : DInt;
      STAT1268 : DInt;
      STAT1269 : DInt;
      STAT1270 : DInt;
      STAT1271 : DInt;
      STAT1272 : DInt;
      STAT1273 : Int;
      STAT1274 : Int := 91;
      STAT1275 : String[10];
      STAT1276 : DInt;
      STAT1277 : DInt;
      STAT1278 : DInt;
      STAT1279 : DInt;
      STAT1280 : DInt;
      STAT1281 : DInt;
      STAT1282 : DInt;
      STAT1283 : DInt;
      STAT1284 : DInt;
      STAT1285 : DInt;
      STAT1286 : DInt;
      STAT1287 : Int;
      STAT1288 : Int := 92;
      STAT1289 : String[10];
      STAT1290 : DInt;
      STAT1291 : DInt;
      STAT1292 : DInt;
      STAT1293 : DInt;
      STAT1294 : DInt;
      STAT1295 : DInt;
      STAT1296 : DInt;
      STAT1297 : DInt;
      STAT1298 : DInt;
      STAT1299 : DInt;
      STAT1300 : DInt;
      STAT1301 : Int;
      STAT1302 : Int := 93;
      STAT1303 : String[10];
      STAT1304 : DInt;
      STAT1305 : DInt;
      STAT1306 : DInt;
      STAT1307 : DInt;
      STAT1308 : DInt;
      STAT1309 : DInt;
      STAT1310 : DInt;
      STAT1311 : DInt;
      STAT1312 : DInt;
      STAT1313 : DInt;
      STAT1314 : DInt;
      STAT1315 : Int;
      STAT1316 : Int := 94;
      STAT1317 : String[10];
      STAT1318 : DInt;
      STAT1319 : DInt;
      STAT1320 : DInt;
      STAT1321 : DInt;
      STAT1322 : DInt;
      STAT1323 : DInt;
      STAT1324 : DInt;
      STAT1325 : DInt;
      STAT1326 : DInt;
      STAT1327 : DInt;
      STAT1328 : DInt;
      STAT1329 : Int;
      STAT1330 : Int := 95;
      STAT1331 : String[10];
      STAT1332 : DInt;
      STAT1333 : DInt;
      STAT1334 : DInt;
      STAT1335 : DInt;
      STAT1336 : DInt;
      STAT1337 : DInt;
      STAT1338 : DInt;
      STAT1339 : DInt;
      STAT1340 : DInt;
      STAT1341 : DInt;
      STAT1342 : DInt;
      STAT1343 : Int;
      STAT1344 : Int := 96;
      STAT1345 : String[10];
      STAT1346 : DInt;
      STAT1347 : DInt;
      STAT1348 : DInt;
      STAT1349 : DInt;
      STAT1350 : DInt;
      STAT1351 : DInt;
      STAT1352 : DInt;
      STAT1353 : DInt;
      STAT1354 : DInt;
      STAT1355 : DInt;
      STAT1356 : DInt;
      STAT1357 : Int;
      STAT1358 : Int := 97;
      STAT1359 : String[10];
      STAT1360 : DInt;
      STAT1361 : DInt;
      STAT1362 : DInt;
      STAT1363 : DInt;
      STAT1364 : DInt;
      STAT1365 : DInt;
      STAT1366 : DInt;
      STAT1367 : DInt;
      STAT1368 : DInt;
      STAT1369 : DInt;
      STAT1370 : DInt;
      STAT1371 : Int;
      STAT1372 : Int := 98;
      STAT1373 : String[10];
      STAT1374 : DInt;
      STAT1375 : DInt;
      STAT1376 : DInt;
      STAT1377 : DInt;
      STAT1378 : DInt;
      STAT1379 : DInt;
      STAT1380 : DInt;
      STAT1381 : DInt;
      STAT1382 : DInt;
      STAT1383 : DInt;
      STAT1384 : DInt;
      STAT1385 : Int;
      STAT1386 : Int := 99;
      STAT1387 : String[10];
      STAT1388 : DInt;
      STAT1389 : DInt;
      STAT1390 : DInt;
      STAT1391 : DInt;
      STAT1392 : DInt;
      STAT1393 : DInt;
      STAT1394 : DInt;
      STAT1395 : DInt;
      STAT1396 : DInt;
      STAT1397 : DInt;
      STAT1398 : DInt;
      STAT1399 : Int;
      STAT1400 : Int := 100;
      STAT1401 : String[10];
      STAT1402 : DInt;
      STAT1403 : DInt;
      STAT1404 : DInt;
      STAT1405 : DInt;
      STAT1406 : DInt;
      STAT1407 : DInt;
      STAT1408 : DInt;
      STAT1409 : DInt;
      STAT1410 : DInt;
      STAT1411 : DInt;
      STAT1412 : DInt;
      STAT1413 : Int;
      STAT1414 : Int := 100;
      STAT1415 : String[10];
      STAT1416 : DInt;
      STAT1417 : DInt;
      STAT1418 : DInt;
      STAT1419 : DInt;
      STAT1420 : DInt;
      STAT1421 : DInt;
      STAT1422 : DInt;
      STAT1423 : DInt;
      STAT1424 : DInt;
      STAT1425 : DInt;
      STAT1426 : DInt;
      STAT1427 : Int;
      STAT1428 : Int := 100;
      STAT1429 : String[10];
      STAT1430 : DInt;
      STAT1431 : DInt;
      STAT1432 : DInt;
      STAT1433 : DInt;
      STAT1434 : DInt;
      STAT1435 : DInt;
      STAT1436 : DInt;
      STAT1437 : DInt;
      STAT1438 : DInt;
      STAT1439 : DInt;
      STAT1440 : DInt;
      STAT1441 : Int;
      STAT1442 : Int := 100;
      STAT1443 : String[10];
      STAT1444 : DInt;
      STAT1445 : DInt;
      STAT1446 : DInt;
      STAT1447 : DInt;
      STAT1448 : DInt;
      STAT1449 : DInt;
      STAT1450 : DInt;
      STAT1451 : DInt;
      STAT1452 : DInt;
      STAT1453 : DInt;
      STAT1454 : DInt;
      STAT1455 : Int;
      STAT1456 : Int := 100;
      STAT1457 : String[10];
      STAT1458 : DInt;
      STAT1459 : DInt;
      STAT1460 : DInt;
      STAT1461 : DInt;
      STAT1462 : DInt;
      STAT1463 : DInt;
      STAT1464 : DInt;
      STAT1465 : DInt;
      STAT1466 : DInt;
      STAT1467 : DInt;
      STAT1468 : DInt;
      STAT1469 : Int;
      STAT1470 : Int := 100;
      STAT1471 : String[10];
      STAT1472 : DInt;
      STAT1473 : DInt;
      STAT1474 : DInt;
      STAT1475 : DInt;
      STAT1476 : DInt;
      STAT1477 : DInt;
      STAT1478 : DInt;
      STAT1479 : DInt;
      STAT1480 : DInt;
      STAT1481 : DInt;
      STAT1482 : DInt;
      STAT1483 : Int;
      STAT1484 : Int := 100;
      STAT1485 : String[10];
      STAT1486 : DInt;
      STAT1487 : DInt;
      STAT1488 : DInt;
      STAT1489 : DInt;
      STAT1490 : DInt;
      STAT1491 : DInt;
      STAT1492 : DInt;
      STAT1493 : DInt;
      STAT1494 : DInt;
      STAT1495 : DInt;
      STAT1496 : DInt;
      STAT1497 : Int;
      STAT1498 : Int := 100;
      STAT1499 : String[10];
      STAT1500 : DInt;
      STAT1501 : DInt;
      STAT1502 : DInt;
      STAT1503 : DInt;
      STAT1504 : DInt;
      STAT1505 : DInt;
      STAT1506 : DInt;
      STAT1507 : DInt;
      STAT1508 : DInt;
      STAT1509 : DInt;
      STAT1510 : DInt;
      STAT1511 : Int;
      STAT1512 : Int := 100;
      STAT1513 : String[10];
      STAT1514 : DInt;
      STAT1515 : DInt;
      STAT1516 : DInt;
      STAT1517 : DInt;
      STAT1518 : DInt;
      STAT1519 : DInt;
      STAT1520 : DInt;
      STAT1521 : DInt;
      STAT1522 : DInt;
      STAT1523 : DInt;
      STAT1524 : DInt;
      STAT1525 : Int;
      STAT1526 : Int := 100;
      STAT1527 : String[10];
      STAT1528 : DInt;
      STAT1529 : DInt;
      STAT1530 : DInt;
      STAT1531 : DInt;
      STAT1532 : DInt;
      STAT1533 : DInt;
      STAT1534 : DInt;
      STAT1535 : DInt;
      STAT1536 : DInt;
      STAT1537 : DInt;
      STAT1538 : DInt;
      STAT1539 : Int;
      STAT1540 : Int := 100;
      STAT1541 : String[10];
      STAT1542 : DInt;
      STAT1543 : DInt;
      STAT1544 : DInt;
      STAT1545 : DInt;
      STAT1546 : DInt;
      STAT1547 : DInt;
      STAT1548 : DInt;
      STAT1549 : DInt;
      STAT1550 : DInt;
      STAT1551 : DInt;
      STAT1552 : DInt;
      STAT1553 : Int;
      STAT1554 : Int := 100;
      STAT1555 : String[10];
      STAT1556 : DInt;
      STAT1557 : DInt;
      STAT1558 : DInt;
      STAT1559 : DInt;
      STAT1560 : DInt;
      STAT1561 : DInt;
      STAT1562 : DInt;
      STAT1563 : DInt;
      STAT1564 : DInt;
      STAT1565 : DInt;
      STAT1566 : DInt;
      STAT1567 : Int;
      STAT1568 : Int := 100;
      STAT1569 : String[10];
      STAT1570 : DInt;
      STAT1571 : DInt;
      STAT1572 : DInt;
      STAT1573 : DInt;
      STAT1574 : DInt;
      STAT1575 : DInt;
      STAT1576 : DInt;
      STAT1577 : DInt;
      STAT1578 : DInt;
      STAT1579 : DInt;
      STAT1580 : DInt;
      STAT1581 : Int;
      STAT1582 : Int := 100;
      STAT1583 : String[10];
      STAT1584 : DInt;
      STAT1585 : DInt;
      STAT1586 : DInt;
      STAT1587 : DInt;
      STAT1588 : DInt;
      STAT1589 : DInt;
      STAT1590 : DInt;
      STAT1591 : DInt;
      STAT1592 : DInt;
      STAT1593 : DInt;
      STAT1594 : DInt;
      STAT1595 : Int;
      STAT1596 : Int := 100;
      STAT1597 : String[10];
      STAT1598 : DInt;
      STAT1599 : DInt;
      STAT1600 : DInt;
      STAT1601 : DInt;
      STAT1602 : DInt;
      STAT1603 : DInt;
      STAT1604 : DInt;
      STAT1605 : DInt;
      STAT1606 : DInt;
      STAT1607 : DInt;
      STAT1608 : DInt;
      STAT1609 : Int;
      STAT1610 : Int := 100;
      STAT1611 : String[10];
      STAT1612 : DInt;
      STAT1613 : DInt;
      STAT1614 : DInt;
      STAT1615 : DInt;
      STAT1616 : DInt;
      STAT1617 : DInt;
      STAT1618 : DInt;
      STAT1619 : DInt;
      STAT1620 : DInt;
      STAT1621 : DInt;
      STAT1622 : DInt;
      STAT1623 : Int;
      STAT1624 : Int := 100;
      STAT1625 : String[10];
      STAT1626 : DInt;
      STAT1627 : DInt;
      STAT1628 : DInt;
      STAT1629 : DInt;
      STAT1630 : DInt;
      STAT1631 : DInt;
      STAT1632 : DInt;
      STAT1633 : DInt;
      STAT1634 : DInt;
      STAT1635 : DInt;
      STAT1636 : DInt;
      STAT1637 : Int;
      STAT1638 : Int := 100;
      STAT1639 : String[10];
      STAT1640 : DInt;
      STAT1641 : DInt;
      STAT1642 : DInt;
      STAT1643 : DInt;
      STAT1644 : DInt;
      STAT1645 : DInt;
      STAT1646 : DInt;
      STAT1647 : DInt;
      STAT1648 : DInt;
      STAT1649 : DInt;
      STAT1650 : DInt;
      STAT1651 : Int;
      STAT1652 : Int := 100;
      STAT1653 : String[10];
      STAT1654 : DInt;
      STAT1655 : DInt;
      STAT1656 : DInt;
      STAT1657 : DInt;
      STAT1658 : DInt;
      STAT1659 : DInt;
      STAT1660 : DInt;
      STAT1661 : DInt;
      STAT1662 : DInt;
      STAT1663 : DInt;
      STAT1664 : DInt;
      STAT1665 : Int;
      STAT1666 : Int := 100;
      STAT1667 : String[10];
      STAT1668 : DInt;
      STAT1669 : DInt;
      STAT1670 : DInt;
      STAT1671 : DInt;
      STAT1672 : DInt;
      STAT1673 : DInt;
      STAT1674 : DInt;
      STAT1675 : DInt;
      STAT1676 : DInt;
      STAT1677 : DInt;
      STAT1678 : DInt;
      STAT1679 : Int;
      STAT1680 : Int := 100;
      STAT1681 : String[10];
      STAT1682 : DInt;
      STAT1683 : DInt;
      STAT1684 : DInt;
      STAT1685 : DInt;
      STAT1686 : DInt;
      STAT1687 : DInt;
      STAT1688 : DInt;
      STAT1689 : DInt;
      STAT1690 : DInt;
      STAT1691 : DInt;
      STAT1692 : DInt;
      STAT1693 : Int;
      STAT1694 : Int := 100;
      STAT1695 : String[10];
      STAT1696 : DInt;
      STAT1697 : DInt;
      STAT1698 : DInt;
      STAT1699 : DInt;
      STAT1700 : DInt;
      STAT1701 : DInt;
      STAT1702 : DInt;
      STAT1703 : DInt;
      STAT1704 : DInt;
      STAT1705 : DInt;
      STAT1706 : DInt;
      STAT1707 : Int;
      STAT1708 : Int := 100;
      STAT1709 : String[10];
      STAT1710 : DInt;
      STAT1711 : DInt;
      STAT1712 : DInt;
      STAT1713 : DInt;
      STAT1714 : DInt;
      STAT1715 : DInt;
      STAT1716 : DInt;
      STAT1717 : DInt;
      STAT1718 : DInt;
      STAT1719 : DInt;
      STAT1720 : DInt;
      STAT1721 : Int;
      STAT1722 : Int := 100;
      STAT1723 : String[10];
      STAT1724 : DInt;
      STAT1725 : DInt;
      STAT1726 : DInt;
      STAT1727 : DInt;
      STAT1728 : DInt;
      STAT1729 : DInt;
      STAT1730 : DInt;
      STAT1731 : DInt;
      STAT1732 : DInt;
      STAT1733 : DInt;
      STAT1734 : DInt;
      STAT1735 : Int;
      STAT1736 : Int := 100;
      STAT1737 : String[10];
      STAT1738 : DInt;
      STAT1739 : DInt;
      STAT1740 : DInt;
      STAT1741 : DInt;
      STAT1742 : DInt;
      STAT1743 : DInt;
      STAT1744 : DInt;
      STAT1745 : DInt;
      STAT1746 : DInt;
      STAT1747 : DInt;
      STAT1748 : DInt;
      STAT1749 : Int;
      STAT1750 : Int := 100;
      STAT1751 : String[10];
      STAT1752 : DInt;
      STAT1753 : DInt;
      STAT1754 : DInt;
      STAT1755 : DInt;
      STAT1756 : DInt;
      STAT1757 : DInt;
      STAT1758 : DInt;
      STAT1759 : DInt;
      STAT1760 : DInt;
      STAT1761 : DInt;
      STAT1762 : DInt;
      STAT1763 : Int;
      STAT1764 : Int := 100;
      STAT1765 : String[10];
      STAT1766 : DInt;
      STAT1767 : DInt;
      STAT1768 : DInt;
      STAT1769 : DInt;
      STAT1770 : DInt;
      STAT1771 : DInt;
      STAT1772 : DInt;
      STAT1773 : DInt;
      STAT1774 : DInt;
      STAT1775 : DInt;
      STAT1776 : DInt;
      STAT1777 : Int;
      STAT1778 : Int := 100;
      STAT1779 : String[10];
      STAT1780 : DInt;
      STAT1781 : DInt;
      STAT1782 : DInt;
      STAT1783 : DInt;
      STAT1784 : DInt;
      STAT1785 : DInt;
      STAT1786 : DInt;
      STAT1787 : DInt;
      STAT1788 : DInt;
      STAT1789 : DInt;
      STAT1790 : DInt;
      STAT1791 : Int;
      STAT1792 : Int := 100;
      STAT1793 : String[10];
      STAT1794 : DInt;
      STAT1795 : DInt;
      STAT1796 : DInt;
      STAT1797 : DInt;
      STAT1798 : DInt;
      STAT1799 : DInt;
      STAT1800 : DInt;
      STAT1801 : DInt;
      STAT1802 : DInt;
      STAT1803 : DInt;
      STAT1804 : DInt;
      STAT1805 : Int;
      STAT1806 : Int := 100;
      STAT1807 : String[10];
      STAT1808 : DInt;
      STAT1809 : DInt;
      STAT1810 : DInt;
      STAT1811 : DInt;
      STAT1812 : DInt;
      STAT1813 : DInt;
      STAT1814 : DInt;
      STAT1815 : DInt;
      STAT1816 : DInt;
      STAT1817 : DInt;
      STAT1818 : DInt;
      STAT1819 : Int;
      STAT1820 : Int := 100;
      STAT1821 : String[10];
      STAT1822 : DInt;
      STAT1823 : DInt;
      STAT1824 : DInt;
      STAT1825 : DInt;
      STAT1826 : DInt;
      STAT1827 : DInt;
      STAT1828 : DInt;
      STAT1829 : DInt;
      STAT1830 : DInt;
      STAT1831 : DInt;
      STAT1832 : DInt;
      STAT1833 : Int;
      STAT1834 : Int := 100;
      STAT1835 : String[10];
      STAT1836 : DInt;
      STAT1837 : DInt;
      STAT1838 : DInt;
      STAT1839 : DInt;
      STAT1840 : DInt;
      STAT1841 : DInt;
      STAT1842 : DInt;
      STAT1843 : DInt;
      STAT1844 : DInt;
      STAT1845 : DInt;
      STAT1846 : DInt;
      STAT1847 : Int;
      STAT1848 : Int := 100;
      STAT1849 : String[10];
      STAT1850 : DInt;
      STAT1851 : DInt;
      STAT1852 : DInt;
      STAT1853 : DInt;
      STAT1854 : DInt;
      STAT1855 : DInt;
      STAT1856 : DInt;
      STAT1857 : DInt;
      STAT1858 : DInt;
      STAT1859 : DInt;
      STAT1860 : DInt;
      STAT1861 : Int;
      STAT1862 : Int := 100;
      STAT1863 : String[10];
      STAT1864 : DInt;
      STAT1865 : DInt;
      STAT1866 : DInt;
      STAT1867 : DInt;
      STAT1868 : DInt;
      STAT1869 : DInt;
      STAT1870 : DInt;
      STAT1871 : DInt;
      STAT1872 : DInt;
      STAT1873 : DInt;
      STAT1874 : DInt;
      STAT1875 : Int;
      STAT1876 : Int := 100;
      STAT1877 : String[10];
      STAT1878 : DInt;
      STAT1879 : DInt;
      STAT1880 : DInt;
      STAT1881 : DInt;
      STAT1882 : DInt;
      STAT1883 : DInt;
      STAT1884 : DInt;
      STAT1885 : DInt;
      STAT1886 : DInt;
      STAT1887 : DInt;
      STAT1888 : DInt;
      STAT1889 : Int;
      STAT1890 : Int := 100;
      STAT1891 : String[10];
      STAT1892 : DInt;
      STAT1893 : DInt;
      STAT1894 : DInt;
      STAT1895 : DInt;
      STAT1896 : DInt;
      STAT1897 : DInt;
      STAT1898 : DInt;
      STAT1899 : DInt;
      STAT1900 : DInt;
      STAT1901 : DInt;
      STAT1902 : DInt;
      STAT1903 : Int;
      STAT1904 : Int := 100;
      STAT1905 : String[10];
      STAT1906 : DInt;
      STAT1907 : DInt;
      STAT1908 : DInt;
      STAT1909 : DInt;
      STAT1910 : DInt;
      STAT1911 : DInt;
      STAT1912 : DInt;
      STAT1913 : DInt;
      STAT1914 : DInt;
      STAT1915 : DInt;
      STAT1916 : DInt;
      STAT1917 : Int;
      STAT1918 : Int := 100;
      STAT1919 : String[10];
      STAT1920 : DInt;
      STAT1921 : DInt;
      STAT1922 : DInt;
      STAT1923 : DInt;
      STAT1924 : DInt;
      STAT1925 : DInt;
      STAT1926 : DInt;
      STAT1927 : DInt;
      STAT1928 : DInt;
      STAT1929 : DInt;
      STAT1930 : DInt;
      STAT1931 : Int;
      STAT1932 : Int := 100;
      STAT1933 : String[10];
      STAT1934 : DInt;
      STAT1935 : DInt;
      STAT1936 : DInt;
      STAT1937 : DInt;
      STAT1938 : DInt;
      STAT1939 : DInt;
      STAT1940 : DInt;
      STAT1941 : DInt;
      STAT1942 : DInt;
      STAT1943 : DInt;
      STAT1944 : DInt;
      STAT1945 : Int;
      STAT1946 : Int := 100;
      STAT1947 : String[10];
      STAT1948 : DInt;
      STAT1949 : DInt;
      STAT1950 : DInt;
      STAT1951 : DInt;
      STAT1952 : DInt;
      STAT1953 : DInt;
      STAT1954 : DInt;
      STAT1955 : DInt;
      STAT1956 : DInt;
      STAT1957 : DInt;
      STAT1958 : DInt;
      STAT1959 : Int;
      STAT1960 : Int := 100;
      STAT1961 : String[10];
      STAT1962 : DInt;
      STAT1963 : DInt;
      STAT1964 : DInt;
      STAT1965 : DInt;
      STAT1966 : DInt;
      STAT1967 : DInt;
      STAT1968 : DInt;
      STAT1969 : DInt;
      STAT1970 : DInt;
      STAT1971 : DInt;
      STAT1972 : DInt;
      STAT1973 : Int;
      STAT1974 : Int := 100;
      STAT1975 : String[10];
      STAT1976 : DInt;
      STAT1977 : DInt;
      STAT1978 : DInt;
      STAT1979 : DInt;
      STAT1980 : DInt;
      STAT1981 : DInt;
      STAT1982 : DInt;
      STAT1983 : DInt;
      STAT1984 : DInt;
      STAT1985 : DInt;
      STAT1986 : DInt;
      STAT1987 : Int;
      STAT1988 : Int := 100;
      STAT1989 : String[10];
      STAT1990 : DInt;
      STAT1991 : DInt;
      STAT1992 : DInt;
      STAT1993 : DInt;
      STAT1994 : DInt;
      STAT1995 : DInt;
      STAT1996 : DInt;
      STAT1997 : DInt;
      STAT1998 : DInt;
      STAT1999 : DInt;
      STAT2000 : DInt;
      STAT2001 : Int;
      STAT2002 : Int := 100;
      STAT2003 : String[10];
      STAT2004 : DInt;
      STAT2005 : DInt;
      STAT2006 : DInt;
      STAT2007 : DInt;
      STAT2008 : DInt;
      STAT2009 : DInt;
      STAT2010 : DInt;
      STAT2011 : DInt;
      STAT2012 : DInt;
      STAT2013 : DInt;
      STAT2014 : DInt;
      STAT2015 : Int;
      STAT2016 : Int := 100;
      STAT2017 : String[10];
      STAT2018 : DInt;
      STAT2019 : DInt;
      STAT2020 : DInt;
      STAT2021 : DInt;
      STAT2022 : DInt;
      STAT2023 : DInt;
      STAT2024 : DInt;
      STAT2025 : DInt;
      STAT2026 : DInt;
      STAT2027 : DInt;
      STAT2028 : DInt;
      STAT2029 : Int;
      STAT2030 : Int := 100;
      STAT2031 : String[10];
      STAT2032 : DInt;
      STAT2033 : DInt;
      STAT2034 : DInt;
      STAT2035 : DInt;
      STAT2036 : DInt;
      STAT2037 : DInt;